REGION Network 8
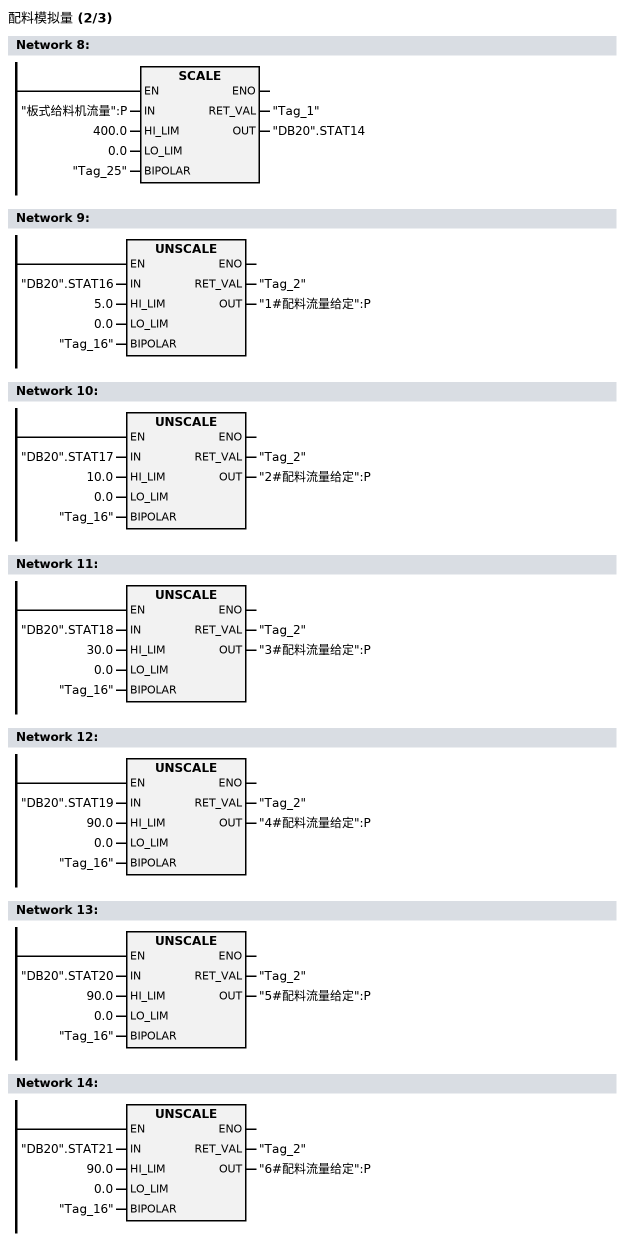
   "Tag_1" := SCALE(IN := "板式给料机流量":P,
                    HI_LIM := 400.0,
                    LO_LIM := 0.0,
                    BIPOLAR := "Tag_25",
                    OUT => "DB20".STAT14);
END_REGION

REGION Network 9
   "Tag_2" := UNSCALE(IN := "DB20".STAT16,
                      HI_LIM := 5.0,
                      LO_LIM := 0.0,
                      BIPOLAR := "Tag_16",
                      OUT => "1#配料流量给定":P);
END_REGION

REGION Network 10
   "Tag_2" := UNSCALE(IN := "DB20".STAT17,
                      HI_LIM := 10.0,
                      LO_LIM := 0.0,
                      BIPOLAR := "Tag_16",
                      OUT => "2#配料流量给定":P);
END_REGION

REGION Network 11
   "Tag_2" := UNSCALE(IN := "DB20".STAT18,
                      HI_LIM := 30.0,
                      LO_LIM := 0.0,
                      BIPOLAR := "Tag_16",
                      OUT => "3#配料流量给定":P);
END_REGION

REGION Network 12
   "Tag_2" := UNSCALE(IN := "DB20".STAT19,
                      HI_LIM := 90.0,
                      LO_LIM := 0.0,
                      BIPOLAR := "Tag_16",
                      OUT => "4#配料流量给定":P);
END_REGION

REGION Network 13
   "Tag_2" := UNSCALE(IN := "DB20".STAT20,
                      HI_LIM := 90.0,
                      LO_LIM := 0.0,
                      BIPOLAR := "Tag_16",
                      OUT => "5#配料流量给定":P);
END_REGION

REGION Network 14
   "Tag_2" := UNSCALE(IN := "DB20".STAT21,
                      HI_LIM := 90.0,
                      LO_LIM := 0.0,
                      BIPOLAR := "Tag_16",
                      OUT => "6#配料流量给定":P);
END_REGION

REGION Network 15
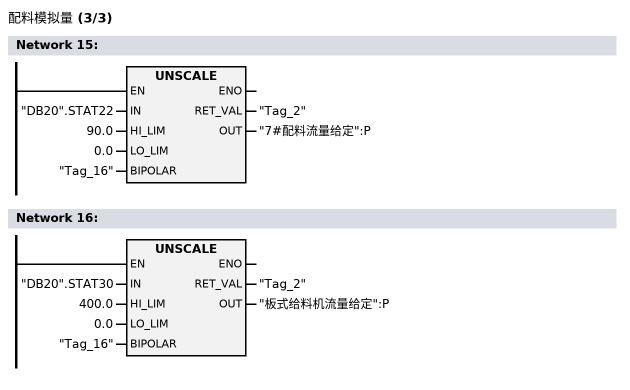
   "Tag_2" := UNSCALE(IN := "DB20".STAT22,
                      HI_LIM := 90.0,
                      LO_LIM := 0.0,
                      BIPOLAR := "Tag_16",
                      OUT => "7#配料流量给定":P);
END_REGION

REGION Network 16
   "Tag_2" := UNSCALE(IN := "DB20".STAT30,
                      HI_LIM := 400.0,
                      LO_LIM := 0.0,
                      BIPOLAR := "Tag_16",
                      OUT => "板式给料机流量给定":P);
END_REGION
END_FUNCTION

FUNCTION "配料累计" : Void   // FC23, LAD
{ S7_Optimized_Access := 'FALSE' }
VERSION : 0.1
   VAR_TEMP   // added for the SCL form of the ladder/FBD networks
      _w1 : Bool;
   END_VAR
BEGIN

REGION Network 1
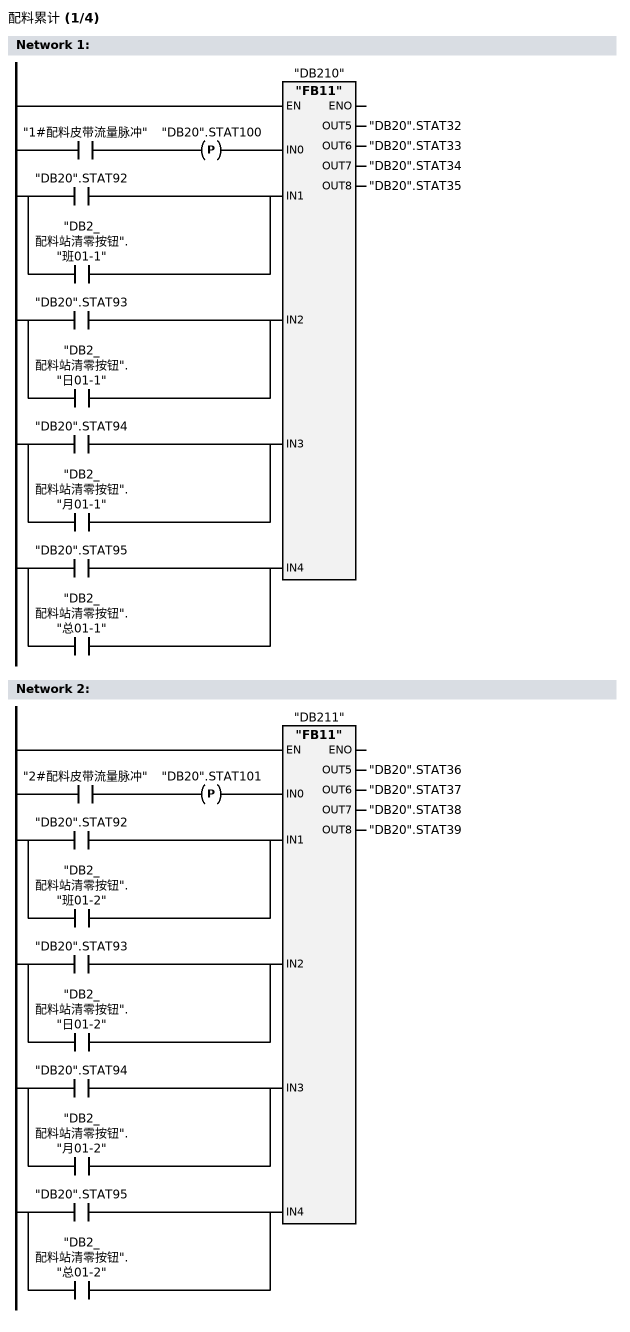
   RUNG wire#powerrail
      "DB210"(IN0 := wire#w1, IN1 := wire#w2, IN2 := wire#w3, IN3 := wire#w4, IN4 := wire#w5, OUT5 => "DB20".STAT32, OUT6 => "DB20".STAT33, OUT7 => "DB20".STAT34, OUT8 => "DB20".STAT35)
   END_RUNG
   RUNG wire#powerrail
      Contact( "1#配料皮带流量脉冲" )
      P_Trig( "DB20".STAT100 )
   END_RUNG wire#w1
   RUNG wire#powerrail
      Contact( "DB20".STAT92 )
   END_RUNG wire#w2
   RUNG wire#powerrail
      Contact( "DB2_配料站清零按钮"."班01-1" )
   END_RUNG wire#w2
   RUNG wire#powerrail
      Contact( "DB20".STAT93 )
   END_RUNG wire#w3
   RUNG wire#powerrail
      Contact( "DB2_配料站清零按钮"."日01-1" )
   END_RUNG wire#w3
   RUNG wire#powerrail
      Contact( "DB20".STAT94 )
   END_RUNG wire#w4
   RUNG wire#powerrail
      Contact( "DB2_配料站清零按钮"."月01-1" )
   END_RUNG wire#w4
   RUNG wire#powerrail
      Contact( "DB20".STAT95 )
   END_RUNG wire#w5
   RUNG wire#powerrail
      Contact( "DB2_配料站清零按钮"."总01-1" )
   END_RUNG wire#w5
   // the same network as SCL:
   #_w1 := "1#配料皮带流量脉冲" AND NOT "DB20".STAT100;   // rising edge
   "DB20".STAT100 := "1#配料皮带流量脉冲";
   "DB210"(IN0 := #_w1,   // "FB11"
           IN1 := "DB20".STAT92 OR "DB2_配料站清零按钮"."班01-1",
           IN2 := "DB20".STAT93 OR "DB2_配料站清零按钮"."日01-1",
           IN3 := "DB20".STAT94 OR "DB2_配料站清零按钮"."月01-1",
           IN4 := "DB20".STAT95 OR "DB2_配料站清零按钮"."总01-1",
           OUT5 => "DB20".STAT32,
           OUT6 => "DB20".STAT33,
           OUT7 => "DB20".STAT34,
           OUT8 => "DB20".STAT35);
END_REGION

REGION Network 2
   RUNG wire#powerrail
      "DB211"(IN0 := wire#w1, IN1 := wire#w2, IN2 := wire#w3, IN3 := wire#w4, IN4 := wire#w5, OUT5 => "DB20".STAT36, OUT6 => "DB20".STAT37, OUT7 => "DB20".STAT38, OUT8 => "DB20".STAT39)
   END_RUNG
   RUNG wire#powerrail
      Contact( "2#配料皮带流量脉冲" )
      P_Trig( "DB20".STAT101 )
   END_RUNG wire#w1
   RUNG wire#powerrail
      Contact( "DB20".STAT92 )
   END_RUNG wire#w2
   RUNG wire#powerrail
      Contact( "DB2_配料站清零按钮"."班01-2" )
   END_RUNG wire#w2
   RUNG wire#powerrail
      Contact( "DB20".STAT93 )
   END_RUNG wire#w3
   RUNG wire#powerrail
      Contact( "DB2_配料站清零按钮"."日01-2" )
   END_RUNG wire#w3
   RUNG wire#powerrail
      Contact( "DB20".STAT94 )
   END_RUNG wire#w4
   RUNG wire#powerrail
      Contact( "DB2_配料站清零按钮"."月01-2" )
   END_RUNG wire#w4
   RUNG wire#powerrail
      Contact( "DB20".STAT95 )
   END_RUNG wire#w5
   RUNG wire#powerrail
      Contact( "DB2_配料站清零按钮"."总01-2" )
   END_RUNG wire#w5
   // the same network as SCL:
   #_w1 := "2#配料皮带流量脉冲" AND NOT "DB20".STAT101;   // rising edge
   "DB20".STAT101 := "2#配料皮带流量脉冲";
   "DB211"(IN0 := #_w1,   // "FB11"
           IN1 := "DB20".STAT92 OR "DB2_配料站清零按钮"."班01-2",
           IN2 := "DB20".STAT93 OR "DB2_配料站清零按钮"."日01-2",
           IN3 := "DB20".STAT94 OR "DB2_配料站清零按钮"."月01-2",
           IN4 := "DB20".STAT95 OR "DB2_配料站清零按钮"."总01-2",
           OUT5 => "DB20".STAT36,
           OUT6 => "DB20".STAT37,
           OUT7 => "DB20".STAT38,
           OUT8 => "DB20".STAT39);
END_REGION

REGION Network 3
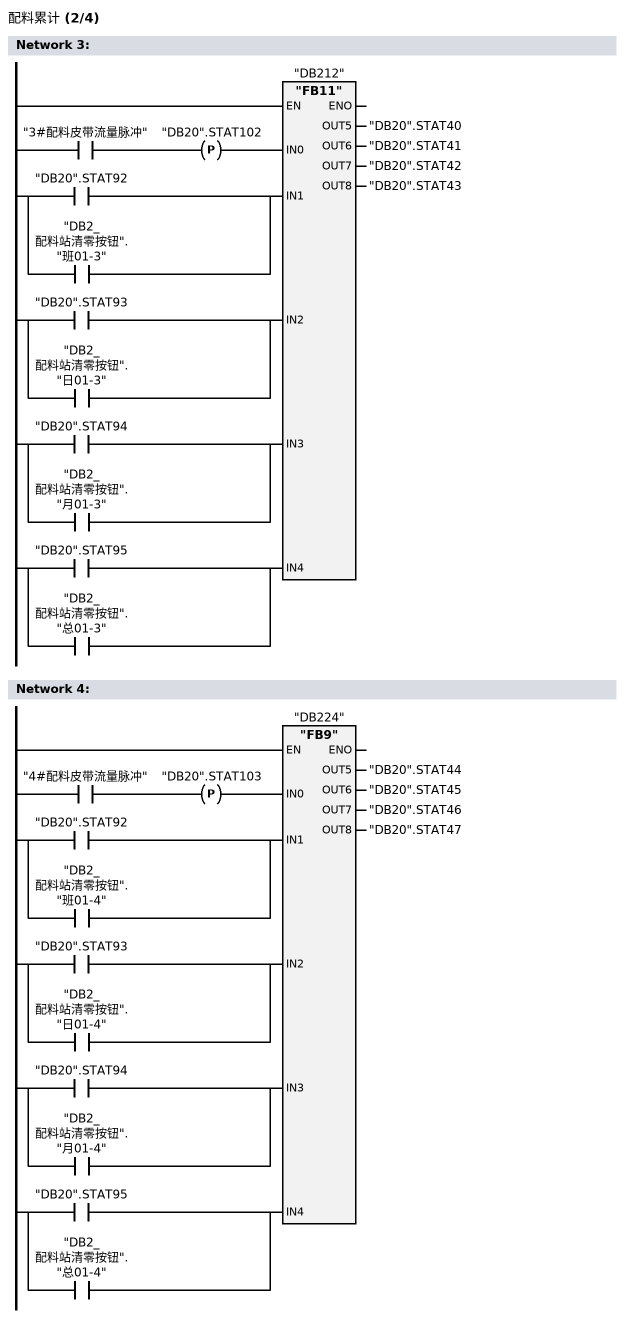
   RUNG wire#powerrail
      "DB212"(IN0 := wire#w1, IN1 := wire#w2, IN2 := wire#w3, IN3 := wire#w4, IN4 := wire#w5, OUT5 => "DB20".STAT40, OUT6 => "DB20".STAT41, OUT7 => "DB20".STAT42, OUT8 => "DB20".STAT43)
   END_RUNG
   RUNG wire#powerrail
      Contact( "3#配料皮带流量脉冲" )
      P_Trig( "DB20".STAT102 )
   END_RUNG wire#w1
   RUNG wire#powerrail
      Contact( "DB20".STAT92 )
   END_RUNG wire#w2
   RUNG wire#powerrail
      Contact( "DB2_配料站清零按钮"."班01-3" )
   END_RUNG wire#w2
   RUNG wire#powerrail
      Contact( "DB20".STAT93 )
   END_RUNG wire#w3
   RUNG wire#powerrail
      Contact( "DB2_配料站清零按钮"."日01-3" )
   END_RUNG wire#w3
   RUNG wire#powerrail
      Contact( "DB20".STAT94 )
   END_RUNG wire#w4
   RUNG wire#powerrail
      Contact( "DB2_配料站清零按钮"."月01-3" )
   END_RUNG wire#w4
   RUNG wire#powerrail
      Contact( "DB20".STAT95 )
   END_RUNG wire#w5
   RUNG wire#powerrail
      Contact( "DB2_配料站清零按钮"."总01-3" )
   END_RUNG wire#w5
   // the same network as SCL:
   #_w1 := "3#配料皮带流量脉冲" AND NOT "DB20".STAT102;   // rising edge
   "DB20".STAT102 := "3#配料皮带流量脉冲";
   "DB212"(IN0 := #_w1,   // "FB11"
           IN1 := "DB20".STAT92 OR "DB2_配料站清零按钮"."班01-3",
           IN2 := "DB20".STAT93 OR "DB2_配料站清零按钮"."日01-3",
           IN3 := "DB20".STAT94 OR "DB2_配料站清零按钮"."月01-3",
           IN4 := "DB20".STAT95 OR "DB2_配料站清零按钮"."总01-3",
           OUT5 => "DB20".STAT40,
           OUT6 => "DB20".STAT41,
           OUT7 => "DB20".STAT42,
           OUT8 => "DB20".STAT43);
END_REGION

REGION Network 4
   RUNG wire#powerrail
      "DB224"(IN0 := wire#w1, IN1 := wire#w2, IN2 := wire#w3, IN3 := wire#w4, IN4 := wire#w5, OUT5 => "DB20".STAT44, OUT6 => "DB20".STAT45, OUT7 => "DB20".STAT46, OUT8 => "DB20".STAT47)
   END_RUNG
   RUNG wire#powerrail
      Contact( "4#配料皮带流量脉冲" )
      P_Trig( "DB20".STAT103 )
   END_RUNG wire#w1
   RUNG wire#powerrail
      Contact( "DB20".STAT92 )
   END_RUNG wire#w2
   RUNG wire#powerrail
      Contact( "DB2_配料站清零按钮"."班01-4" )
   END_RUNG wire#w2
   RUNG wire#powerrail
      Contact( "DB20".STAT93 )
   END_RUNG wire#w3
   RUNG wire#powerrail
      Contact( "DB2_配料站清零按钮"."日01-4" )
   END_RUNG wire#w3
   RUNG wire#powerrail
      Contact( "DB20".STAT94 )
   END_RUNG wire#w4
   RUNG wire#powerrail
      Contact( "DB2_配料站清零按钮"."月01-4" )
   END_RUNG wire#w4
   RUNG wire#powerrail
      Contact( "DB20".STAT95 )
   END_RUNG wire#w5
   RUNG wire#powerrail
      Contact( "DB2_配料站清零按钮"."总01-4" )
   END_RUNG wire#w5
   // the same network as SCL:
   #_w1 := "4#配料皮带流量脉冲" AND NOT "DB20".STAT103;   // rising edge
   "DB20".STAT103 := "4#配料皮带流量脉冲";
   "DB224"(IN0 := #_w1,   // "FB9"
           IN1 := "DB20".STAT92 OR "DB2_配料站清零按钮"."班01-4",
           IN2 := "DB20".STAT93 OR "DB2_配料站清零按钮"."日01-4",
           IN3 := "DB20".STAT94 OR "DB2_配料站清零按钮"."月01-4",
           IN4 := "DB20".STAT95 OR "DB2_配料站清零按钮"."总01-4",
           OUT5 => "DB20".STAT44,
           OUT6 => "DB20".STAT45,
           OUT7 => "DB20".STAT46,
           OUT8 => "DB20".STAT47);
END_REGION

REGION Network 5
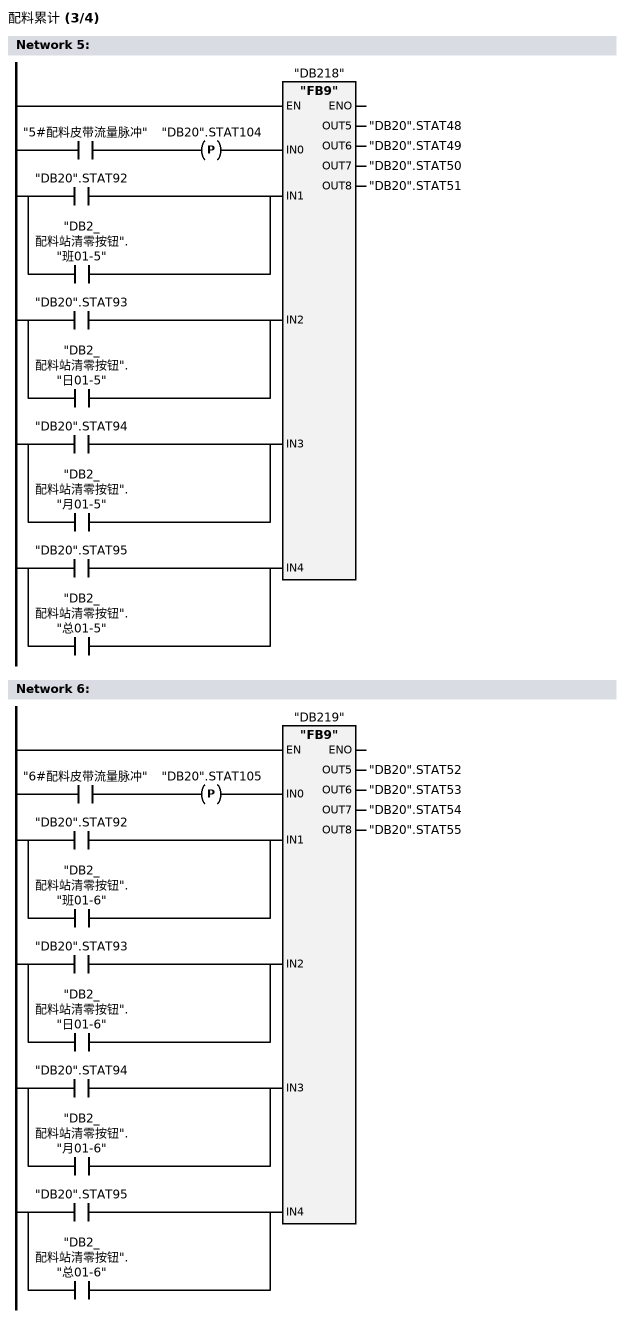
   RUNG wire#powerrail
      "DB218"(IN0 := wire#w1, IN1 := wire#w2, IN2 := wire#w3, IN3 := wire#w4, IN4 := wire#w5, OUT5 => "DB20".STAT48, OUT6 => "DB20".STAT49, OUT7 => "DB20".STAT50, OUT8 => "DB20".STAT51)
   END_RUNG
   RUNG wire#powerrail
      Contact( "5#配料皮带流量脉冲" )
      P_Trig( "DB20".STAT104 )
   END_RUNG wire#w1
   RUNG wire#powerrail
      Contact( "DB20".STAT92 )
   END_RUNG wire#w2
   RUNG wire#powerrail
      Contact( "DB2_配料站清零按钮"."班01-5" )
   END_RUNG wire#w2
   RUNG wire#powerrail
      Contact( "DB20".STAT93 )
   END_RUNG wire#w3
   RUNG wire#powerrail
      Contact( "DB2_配料站清零按钮"."日01-5" )
   END_RUNG wire#w3
   RUNG wire#powerrail
      Contact( "DB20".STAT94 )
   END_RUNG wire#w4
   RUNG wire#powerrail
      Contact( "DB2_配料站清零按钮"."月01-5" )
   END_RUNG wire#w4
   RUNG wire#powerrail
      Contact( "DB20".STAT95 )
   END_RUNG wire#w5
   RUNG wire#powerrail
      Contact( "DB2_配料站清零按钮"."总01-5" )
   END_RUNG wire#w5
   // the same network as SCL:
   #_w1 := "5#配料皮带流量脉冲" AND NOT "DB20".STAT104;   // rising edge
   "DB20".STAT104 := "5#配料皮带流量脉冲";
   "DB218"(IN0 := #_w1,   // "FB9"
           IN1 := "DB20".STAT92 OR "DB2_配料站清零按钮"."班01-5",
           IN2 := "DB20".STAT93 OR "DB2_配料站清零按钮"."日01-5",
           IN3 := "DB20".STAT94 OR "DB2_配料站清零按钮"."月01-5",
           IN4 := "DB20".STAT95 OR "DB2_配料站清零按钮"."总01-5",
           OUT5 => "DB20".STAT48,
           OUT6 => "DB20".STAT49,
           OUT7 => "DB20".STAT50,
           OUT8 => "DB20".STAT51);
END_REGION

REGION Network 6
   RUNG wire#powerrail
      "DB219"(IN0 := wire#w1, IN1 := wire#w2, IN2 := wire#w3, IN3 := wire#w4, IN4 := wire#w5, OUT5 => "DB20".STAT52, OUT6 => "DB20".STAT53, OUT7 => "DB20".STAT54, OUT8 => "DB20".STAT55)
   END_RUNG
   RUNG wire#powerrail
      Contact( "6#配料皮带流量脉冲" )
      P_Trig( "DB20".STAT105 )
   END_RUNG wire#w1
   RUNG wire#powerrail
      Contact( "DB20".STAT92 )
   END_RUNG wire#w2
   RUNG wire#powerrail
      Contact( "DB2_配料站清零按钮"."班01-6" )
   END_RUNG wire#w2
   RUNG wire#powerrail
      Contact( "DB20".STAT93 )
   END_RUNG wire#w3
   RUNG wire#powerrail
      Contact( "DB2_配料站清零按钮"."日01-6" )
   END_RUNG wire#w3
   RUNG wire#powerrail
      Contact( "DB20".STAT94 )
   END_RUNG wire#w4
   RUNG wire#powerrail
      Contact( "DB2_配料站清零按钮"."月01-6" )
   END_RUNG wire#w4
   RUNG wire#powerrail
      Contact( "DB20".STAT95 )
   END_RUNG wire#w5
   RUNG wire#powerrail
      Contact( "DB2_配料站清零按钮"."总01-6" )
   END_RUNG wire#w5
   // the same network as SCL:
   #_w1 := "6#配料皮带流量脉冲" AND NOT "DB20".STAT105;   // rising edge
   "DB20".STAT105 := "6#配料皮带流量脉冲";
   "DB219"(IN0 := #_w1,   // "FB9"
           IN1 := "DB20".STAT92 OR "DB2_配料站清零按钮"."班01-6",
           IN2 := "DB20".STAT93 OR "DB2_配料站清零按钮"."日01-6",
           IN3 := "DB20".STAT94 OR "DB2_配料站清零按钮"."月01-6",
           IN4 := "DB20".STAT95 OR "DB2_配料站清零按钮"."总01-6",
           OUT5 => "DB20".STAT52,
           OUT6 => "DB20".STAT53,
           OUT7 => "DB20".STAT54,
           OUT8 => "DB20".STAT55);
END_REGION

REGION Network 7
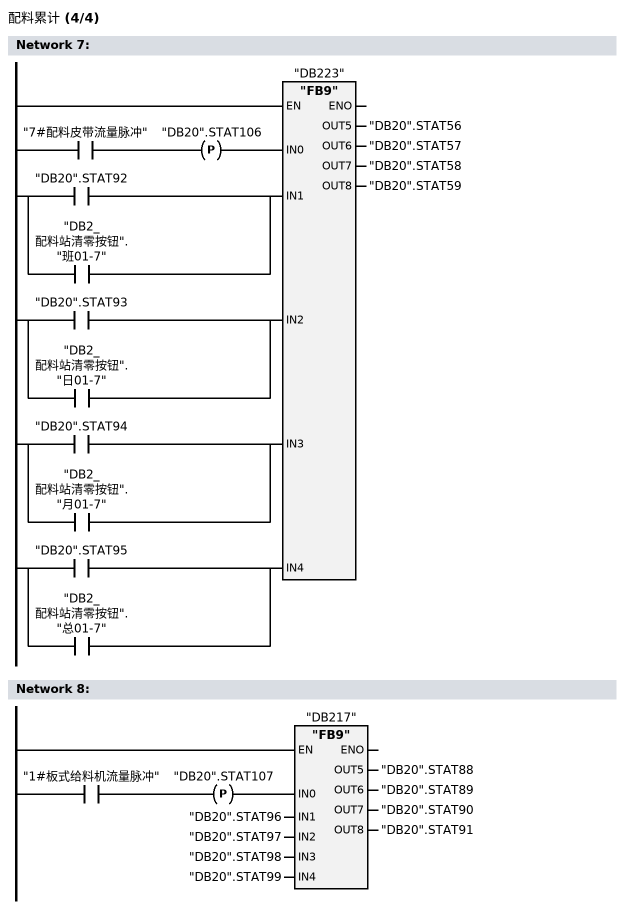
   RUNG wire#powerrail
      "DB223"(IN0 := wire#w1, IN1 := wire#w2, IN2 := wire#w3, IN3 := wire#w4, IN4 := wire#w5, OUT5 => "DB20".STAT56, OUT6 => "DB20".STAT57, OUT7 => "DB20".STAT58, OUT8 => "DB20".STAT59)
   END_RUNG
   RUNG wire#powerrail
      Contact( "7#配料皮带流量脉冲" )
      P_Trig( "DB20".STAT106 )
   END_RUNG wire#w1
   RUNG wire#powerrail
      Contact( "DB20".STAT92 )
   END_RUNG wire#w2
   RUNG wire#powerrail
      Contact( "DB2_配料站清零按钮"."班01-7" )
   END_RUNG wire#w2
   RUNG wire#powerrail
      Contact( "DB20".STAT93 )
   END_RUNG wire#w3
   RUNG wire#powerrail
      Contact( "DB2_配料站清零按钮"."日01-7" )
   END_RUNG wire#w3
   RUNG wire#powerrail
      Contact( "DB20".STAT94 )
   END_RUNG wire#w4
   RUNG wire#powerrail
      Contact( "DB2_配料站清零按钮"."月01-7" )
   END_RUNG wire#w4
   RUNG wire#powerrail
      Contact( "DB20".STAT95 )
   END_RUNG wire#w5
   RUNG wire#powerrail
      Contact( "DB2_配料站清零按钮"."总01-7" )
   END_RUNG wire#w5
   // the same network as SCL:
   #_w1 := "7#配料皮带流量脉冲" AND NOT "DB20".STAT106;   // rising edge
   "DB20".STAT106 := "7#配料皮带流量脉冲";
   "DB223"(IN0 := #_w1,   // "FB9"
           IN1 := "DB20".STAT92 OR "DB2_配料站清零按钮"."班01-7",
           IN2 := "DB20".STAT93 OR "DB2_配料站清零按钮"."日01-7",
           IN3 := "DB20".STAT94 OR "DB2_配料站清零按钮"."月01-7",
           IN4 := "DB20".STAT95 OR "DB2_配料站清零按钮"."总01-7",
           OUT5 => "DB20".STAT56,
           OUT6 => "DB20".STAT57,
           OUT7 => "DB20".STAT58,
           OUT8 => "DB20".STAT59);
END_REGION

REGION Network 8
   RUNG wire#powerrail
      "DB217"(IN0 := wire#w1, IN1 := "DB20".STAT96, IN2 := "DB20".STAT97, IN3 := "DB20".STAT98, IN4 := "DB20".STAT99, OUT5 => "DB20".STAT88, OUT6 => "DB20".STAT89, OUT7 => "DB20".STAT90, OUT8 => "DB20".STAT91)
   END_RUNG
   RUNG wire#powerrail
      Contact( "1#板式给料机流量脉冲" )
      P_Trig( "DB20".STAT107 )
   END_RUNG wire#w1
   // the same network as SCL:
   #_w1 := "1#板式给料机流量脉冲" AND NOT "DB20".STAT107;   // rising edge
   "DB20".STAT107 := "1#板式给料机流量脉冲";
   "DB217"(IN0 := #_w1,   // "FB9"
           IN1 := "DB20".STAT96,
           IN2 := "DB20".STAT97,
           IN3 := "DB20".STAT98,
           IN4 := "DB20".STAT99,
           OUT5 => "DB20".STAT88,
           OUT6 => "DB20".STAT89,
           OUT7 => "DB20".STAT90,
           OUT8 => "DB20".STAT91);
END_REGION
END_FUNCTION

FUNCTION "回转窑变频器驱动块" : Void   // FC111, LAD
{ S7_Optimized_Access := 'FALSE' }
VERSION : 0.1
   VAR_INPUT
      IN0 : Bool;   // IN0
      IN1 : Bool;   // IN1
      IN2 : Bool;   // IN2
      IN3 : Bool;   // IN3
      IN4 : Bool;   // IN4
      IN5 : Bool;   // IN5
      IN6 : Bool;   // IN6
      IN7 : Bool;   // IN7
      IN8 : Bool;   // IN8
   END_VAR
   VAR_IN_OUT
      OUT9 : Bool;   // OUT9
   END_VAR
BEGIN

REGION Network 1: OUT9
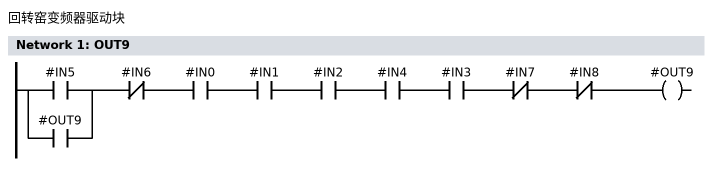
   RUNG wire#powerrail
      Contact( #IN5 )
      wire#w1
      I_Contact( #IN6 )
      Contact( #IN0 )
      Contact( #IN1 )
      Contact( #IN2 )
      Contact( #IN4 )
      Contact( #IN3 )
      I_Contact( #IN7 )
      I_Contact( #IN8 )
      Coil( #OUT9 )
   END_RUNG
   RUNG wire#powerrail
      Contact( #OUT9 )
   END_RUNG wire#w1
   // the same network as SCL:
   #OUT9 := (#IN5 OR #OUT9) AND NOT #IN6 AND #IN0 AND #IN1 AND #IN2 AND #IN4 AND #IN3 AND NOT #IN7 AND NOT #IN8;
END_REGION
END_FUNCTION

FUNCTION "回转窑接触器合闸块" : Void   // FC112, LAD
{ S7_Optimized_Access := 'FALSE' }
VERSION : 0.1
   VAR_INPUT
      IN0 : Bool;   // IN0
      IN1 : Bool;   // IN1
      IN2 : Bool;   // IN2
   END_VAR
   VAR_IN_OUT
      OUT3 : Bool;   // OUT3
   END_VAR
BEGIN

REGION Network 1: OUT3
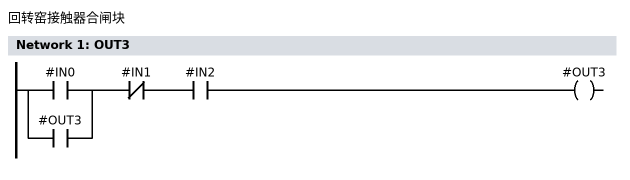
   RUNG wire#powerrail
      Contact( #IN0 )
      wire#w1
      I_Contact( #IN1 )
      Contact( #IN2 )
      Coil( #OUT3 )
   END_RUNG
   RUNG wire#powerrail
      Contact( #OUT3 )
   END_RUNG wire#w1
   // the same network as SCL:
   #OUT3 := (#IN0 OR #OUT3) AND NOT #IN1 AND #IN2;
END_REGION
END_FUNCTION

FUNCTION "稀油站功能块" : Void   // FC113, LAD
{ S7_Optimized_Access := 'FALSE' }
VERSION : 0.1
   VAR_INPUT
      LR1 : Bool;
      FAT1_1 : Bool;
      FAT1_2 : Bool;
      ST1 : Bool;
      STP1 : Bool;
      LR2 : Bool;
      FAT2_1 : Bool;
      FAT2_2 : Bool;
      ST2 : Bool;
      STP2 : Bool;
   END_VAR
   VAR_IN_OUT
      OUT10 : Bool;
      OUT11 : Bool;
   END_VAR
BEGIN

REGION Network 1
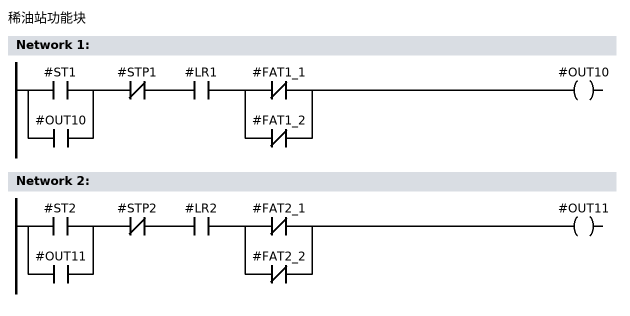
   RUNG wire#powerrail
      Contact( #ST1 )
      wire#w1
      I_Contact( #STP1 )
      Contact( #LR1 )
      wire#w2
      I_Contact( #FAT1_1 )
      wire#w3
      Coil( #OUT10 )
   END_RUNG
   RUNG wire#powerrail
      Contact( #OUT10 )
   END_RUNG wire#w1
   RUNG wire#w2
      I_Contact( #FAT1_2 )
   END_RUNG wire#w3
   // the same network as SCL:
   #OUT10 := (#ST1 OR #OUT10) AND NOT #STP1 AND #LR1 AND (NOT #FAT1_1 OR NOT #FAT1_2);
END_REGION

REGION Network 2
   RUNG wire#powerrail
      Contact( #ST2 )
      wire#w1
      I_Contact( #STP2 )
      Contact( #LR2 )
      wire#w2
      I_Contact( #FAT2_1 )
      wire#w3
      Coil( #OUT11 )
   END_RUNG
   RUNG wire#powerrail
      Contact( #OUT11 )
   END_RUNG wire#w1
   RUNG wire#w2
      I_Contact( #FAT2_2 )
   END_RUNG wire#w3
   // the same network as SCL:
   #OUT11 := (#ST2 OR #OUT11) AND NOT #STP2 AND #LR2 AND (NOT #FAT2_1 OR NOT #FAT2_2);
END_REGION
END_FUNCTION

FUNCTION "电机功能块" : Void   // FC114, LAD
{ S7_Optimized_Access := 'FALSE' }
VERSION : 0.1
   VAR_INPUT
      LR : Bool;
      FAULT : Bool;
      START : Bool;
      STOP : Bool;
   END_VAR
   VAR_IN_OUT
      OUT : Bool;
   END_VAR
BEGIN

REGION Network 1
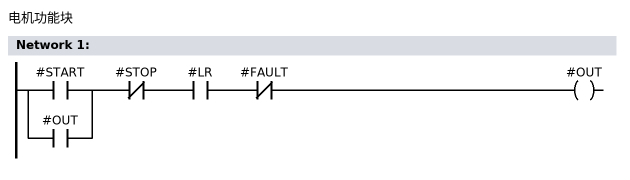
   RUNG wire#powerrail
      Contact( #START )
      wire#w1
      I_Contact( #STOP )
      Contact( #LR )
      I_Contact( #FAULT )
      Coil( #OUT )
   END_RUNG
   RUNG wire#powerrail
      Contact( #OUT )
   END_RUNG wire#w1
   // the same network as SCL:
   #OUT := (#START OR #OUT) AND NOT #STOP AND #LR AND NOT #FAULT;
END_REGION
END_FUNCTION

FUNCTION "皮带功能块" : Void   // FC115, LAD
{ S7_Optimized_Access := 'FALSE' }
VERSION : 0.1
   VAR_INPUT
      LR : Bool;
      FAULT : Bool;
      STOP : Bool;
      IN3 : Bool;
   END_VAR
   VAR_IN_OUT
      OUT : Bool;
   END_VAR
BEGIN

REGION Network 1
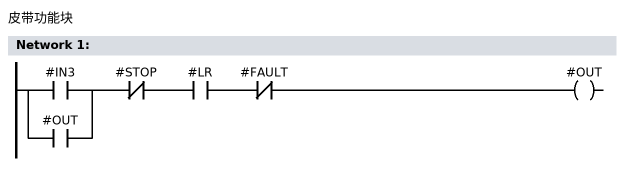
   RUNG wire#powerrail
      Contact( #IN3 )
      wire#w1
      I_Contact( #STOP )
      Contact( #LR )
      I_Contact( #FAULT )
      Coil( #OUT )
   END_RUNG
   RUNG wire#powerrail
      Contact( #OUT )
   END_RUNG wire#w1
   // the same network as SCL:
   #OUT := (#IN3 OR #OUT) AND NOT #STOP AND #LR AND NOT #FAULT;
END_REGION
END_FUNCTION

FUNCTION "脉冲累计功能块" : Void   // FC116, LAD
{ S7_Optimized_Access := 'FALSE' }
VERSION : 0.1
   VAR_INPUT
      IN0 : Bool;
      IN1 : Bool;
   END_VAR
   VAR_OUTPUT
      OUT2 : Real;
   END_VAR
   VAR_TEMP
      TEMP3 : Bool;
      TEMP4 : Real;
      TEMP5 : Real;
      TEMP6 : Real;
   END_VAR
   VAR_TEMP   // added for the SCL form of the ladder/FBD networks
      _w1 : Bool;
   END_VAR
BEGIN

REGION Network 1
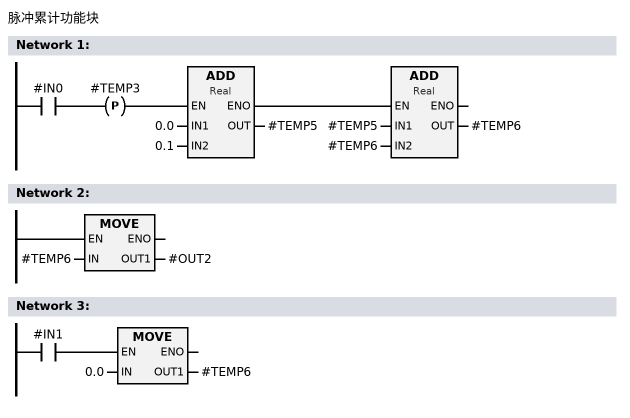
   RUNG wire#powerrail
      Contact( #IN0 )
      P_Trig( #TEMP3 )
      { S7_Templates := "SrcType := Real"; S7_GenerateENO := "TRUE" } Add(in1 := 0.0, in2 := 0.1, out => #TEMP5)
      { S7_Templates := "SrcType := Real"; S7_GenerateENO := "TRUE" } Add(in1 := #TEMP5, in2 := #TEMP6, out => #TEMP6)
   END_RUNG
   // the same network as SCL:
   // ENO of a box is taken as its EN; it also drops when the box reports an error
   #_w1 := #IN0 AND NOT #TEMP3;   // rising edge
   #TEMP3 := #IN0;
   IF #_w1 THEN
       #TEMP5 := 0.0 + 0.1;
       #TEMP6 := #TEMP5 + #TEMP6;
   END_IF;
END_REGION

REGION Network 2
   RUNG wire#powerrail
      { S7_GenerateENO := "TRUE" } Move(in := #TEMP6, out1 => #OUT2)
   END_RUNG
   // the same network as SCL:
   #OUT2 := #TEMP6;
END_REGION

REGION Network 3
   RUNG wire#powerrail
      Contact( #IN1 )
      { S7_GenerateENO := "TRUE" } Move(in := 0.0, out1 => #TEMP6)
   END_RUNG
   // the same network as SCL:
   IF #IN1 THEN #TEMP6 := 0.0; END_IF;
END_REGION

REGION Network 4 (STL)
         SET;
         SAVE;
END_REGION
END_FUNCTION

ORGANIZATION_BLOCK "Main"   // OB1, LAD, ProgramCycle
{ S7_Optimized_Access := 'FALSE' }
VERSION : 0.1
   VAR_TEMP
      TEMP0 : Byte;
      TEMP1 : Byte;
      TEMP2 : Byte;
      TEMP3 : Byte;
      TEMP4 : Byte;
      TEMP5 : Byte;
      TEMP6 : Int;
      TEMP7 : Int;
      TEMP8 : Int;
      TEMP9 : Date_And_Time;
   END_VAR
BEGIN

REGION Network 1